(* Logix 5000 project; controller PLC_MCC1300_75F1 vendor 1 type 14 code 166 rev 32.11; software revision 32.04; part 53 of 83 *)
(* tags used below, declared in another part *)
   AUX_tConvoy_SL_NULL : UDT_Convoy_SL;
   AUX_xInitialize : BOOL;
   CONST_rgdDestMask : DINT[32];   // Destination Mask
   CONST_tPlant : UDT_PLANT_CONSTANTS;
   GP_TrackingGetFirstPlateInConveyor : GP_TrackingGetFirstPlateInConveyor;
   GP_TrackingPresencePlate : GP_TrackingPresencePlate;
   GP_TrackingSearchPlate : GP_TrackingSearchPlate;
   M310_M1_DR_R1 : AXIS_CIP_DRIVE;
   M310_xReqStopPrevConvForPos : BOOL;
   M310Popup : MAC_Popup_ZC[2];
   M310Popup_ReentryCap : UDT_ConvoyCap_ZC;
   M310Popup_SL_DATA : UDT_Convoy_SL;
   M310Popup_xDrivePosEnable : BOOL;
   M310Popup_xEndRise : BOOL;
   M310Popup_xEndRiseWaitingForCondition : BOOL;
   Sbr_INO_tConvoy_SL : UDT_Convoy_SL;
   TMP_d : DINT;
   TMP_dBaryc_ins_max : DINT;
   TMP_dBaryc_ins_min : DINT;
   TMP_dIndex : DINT;
   TMP_dIndex2 : DINT;
   TMP_dIndex3 : DINT;
   TMP_dStart0 : DINT;
   TMP_dStart1 : DINT;
   TMP_dStartSearchStop : DINT;
   TMP_dStop0 : DINT;
   TMP_dStop1 : DINT;
   TMP_dStopSearchStop : DINT;
   TMP_StartPlusLength : DINT;
   TMP_xAllCullet : BOOL;
   TMP_xAllLiteToCullet : BOOL;
   TMP_xAtLeastOneForSideLeg : BOOL;
   TMP_xPosHead : BOOL;
   TMP_xReqStopM310M1 : BOOL;
   TMP_xReqStopM310M2 : BOOL;
   TMP_xReqStopM310M3 : BOOL;
   xAlwaysOFF : BOOL;
   xDebugOFF : BOOL;
   Z300_BufferPlate : UDT_LINE_BUFFER_PLATE;
   Z300_Conveyor : UDT_StandConv[29];
   Z300_Conveyor_IN_MOTION : MAC_Conveyor_ZC_IN_MOTION[29];
   Z300_LineTracking : UDT_LINE_TRACKING;
   Z301 : MAC_Zone_ML;
(* MainProgram, continued *)

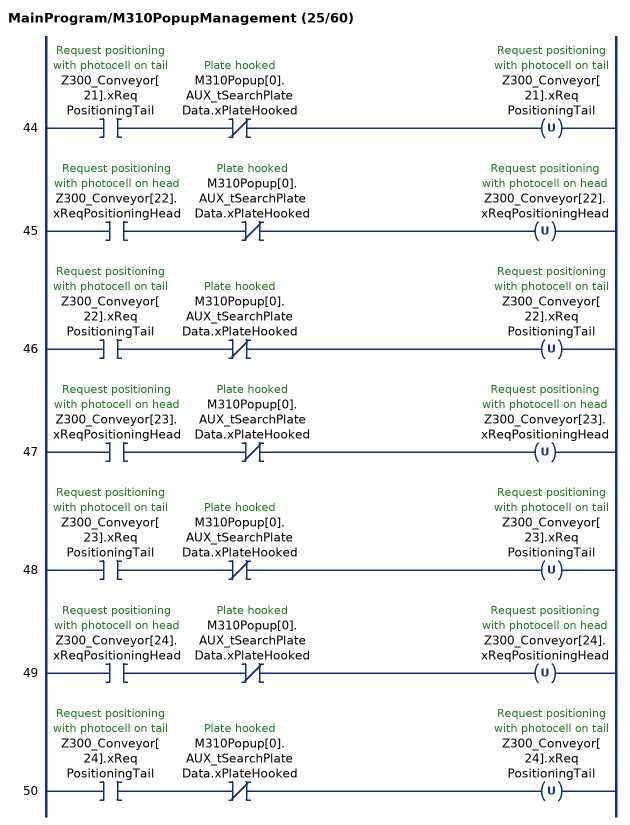
   [picture p841: MainProgram/M310PopupManagement rungs 44-50]
   44: XIC(Z300_Conveyor[21].xReqPositioningTail)XIO(M310Popup[0].AUX_tSearchPlateData.xPlateHooked)OTU(Z300_Conveyor[21].xReqPositioningTail);
   45: XIC(Z300_Conveyor[22].xReqPositioningHead)XIO(M310Popup[0].AUX_tSearchPlateData.xPlateHooked)OTU(Z300_Conveyor[22].xReqPositioningHead);
   46: XIC(Z300_Conveyor[22].xReqPositioningTail)XIO(M310Popup[0].AUX_tSearchPlateData.xPlateHooked)OTU(Z300_Conveyor[22].xReqPositioningTail);
   47: XIC(Z300_Conveyor[23].xReqPositioningHead)XIO(M310Popup[0].AUX_tSearchPlateData.xPlateHooked)OTU(Z300_Conveyor[23].xReqPositioningHead);
   48: XIC(Z300_Conveyor[23].xReqPositioningTail)XIO(M310Popup[0].AUX_tSearchPlateData.xPlateHooked)OTU(Z300_Conveyor[23].xReqPositioningTail);
   49: XIC(Z300_Conveyor[24].xReqPositioningHead)XIO(M310Popup[0].AUX_tSearchPlateData.xPlateHooked)OTU(Z300_Conveyor[24].xReqPositioningHead);
   50: XIC(Z300_Conveyor[24].xReqPositioningTail)XIO(M310Popup[0].AUX_tSearchPlateData.xPlateHooked)OTU(Z300_Conveyor[24].xReqPositioningTail);
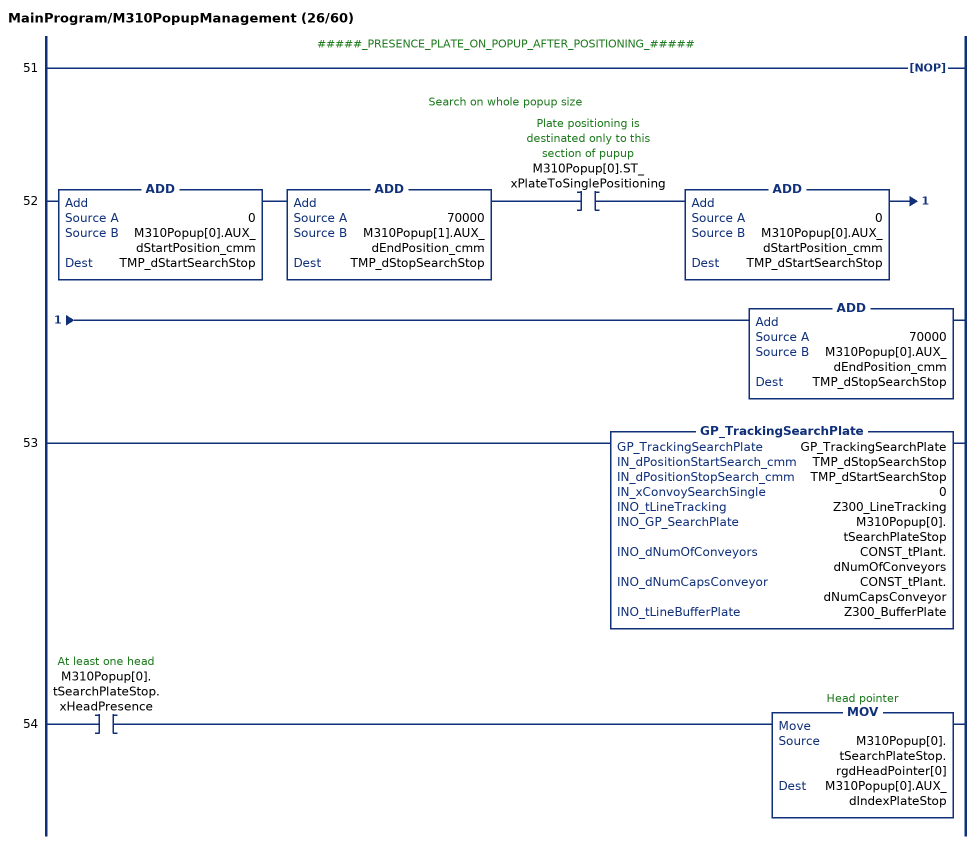
   // #####_PRESENCE_PLATE_ON_POPUP_AFTER_POSITIONING_#####
   51: NOP();
   // Search on whole popup size
   52: ADD(0,M310Popup[0].AUX_dStartPosition_cmm,TMP_dStartSearchStop)ADD(70000,M310Popup[1].AUX_dEndPosition_cmm,TMP_dStopSearchStop)XIC(M310Popup[0].ST_xPlateToSinglePositioning)ADD(0,M310Popup[0].AUX_dStartPosition_cmm,TMP_dStartSearchStop)ADD(70000,M310Popup[0].AUX_dEndPosition_cmm,TMP_dStopSearchStop);
   53: GP_TrackingSearchPlate(GP_TrackingSearchPlate,TMP_dStopSearchStop,TMP_dStartSearchStop,0,Z300_LineTracking,M310Popup[0].tSearchPlateStop,CONST_tPlant.dNumOfConveyors,CONST_tPlant.dNumCapsConveyor,Z300_BufferPlate);
   54: XIC(M310Popup[0].tSearchPlateStop.xHeadPresence)MOV(M310Popup[0].tSearchPlateStop.rgdHeadPointer[0],M310Popup[0].AUX_dIndexPlateStop);
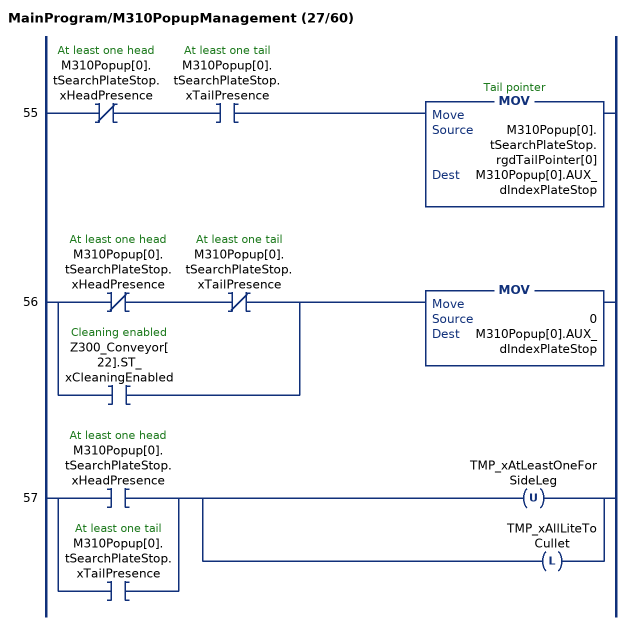
   55: XIO(M310Popup[0].tSearchPlateStop.xHeadPresence)XIC(M310Popup[0].tSearchPlateStop.xTailPresence)MOV(M310Popup[0].tSearchPlateStop.rgdTailPointer[0],M310Popup[0].AUX_dIndexPlateStop);
   56: [XIO(M310Popup[0].tSearchPlateStop.xHeadPresence) XIO(M310Popup[0].tSearchPlateStop.xTailPresence) ,XIC(Z300_Conveyor[22].ST_xCleaningEnabled) ]MOV(0,M310Popup[0].AUX_dIndexPlateStop);
   57: [XIC(M310Popup[0].tSearchPlateStop.xHeadPresence) ,XIC(M310Popup[0].tSearchPlateStop.xTailPresence) ][OTU(TMP_xAtLeastOneForSideLeg) ,OTL(TMP_xAllLiteToCullet) ];
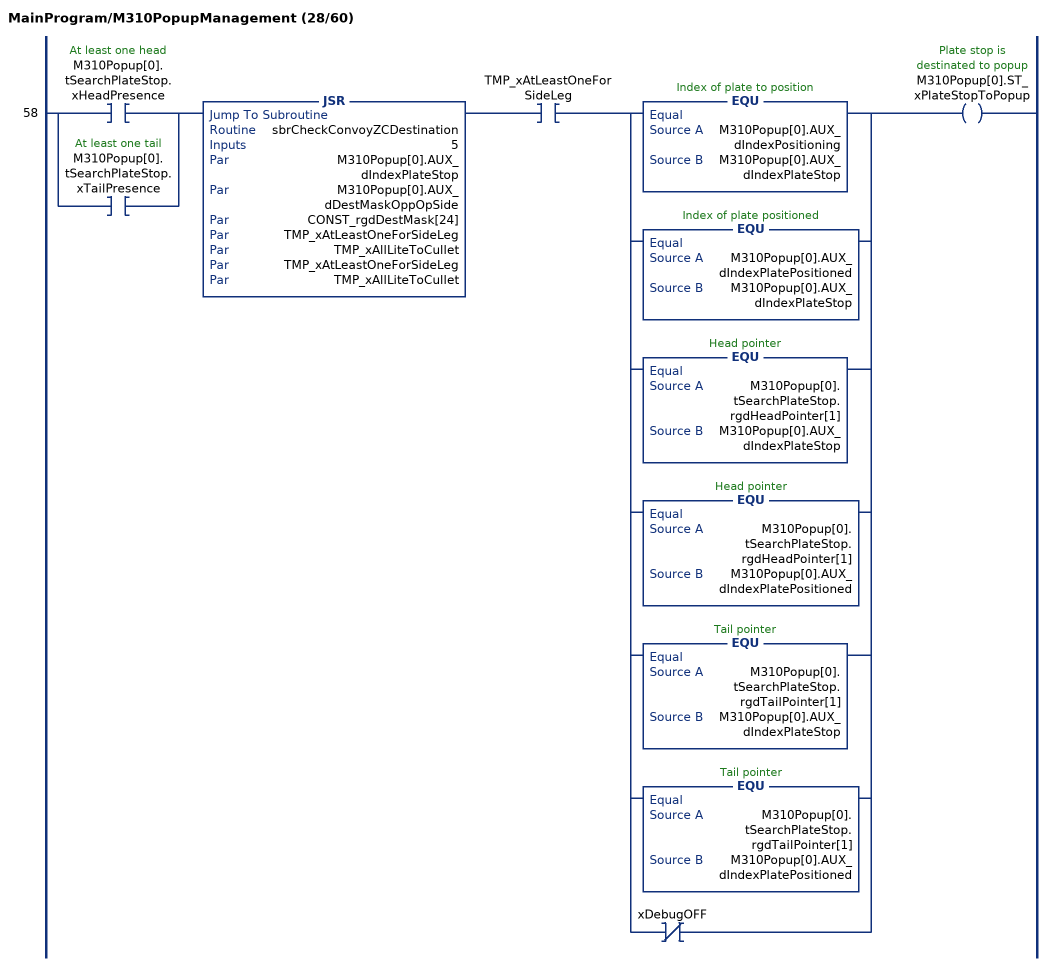
   58: [XIC(M310Popup[0].tSearchPlateStop.xHeadPresence) ,XIC(M310Popup[0].tSearchPlateStop.xTailPresence) ]JSR(sbrCheckConvoyZCDestination,5,M310Popup[0].AUX_dIndexPlateStop,M310Popup[0].AUX_dDestMaskOppOpSide,CONST_rgdDestMask[24],TMP_xAtLeastOneForSideLeg,TMP_xAllLiteToCullet,TMP_xAtLeastOneForSideLeg,TMP_xAllLiteToCullet)XIC(TMP_xAtLeastOneForSideLeg)[EQU(M310Popup[0].AUX_dIndexPositioning,M310Popup[0].AUX_dIndexPlateStop) ,EQU(M310Popup[0].AUX_dIndexPlatePositioned,M310Popup[0].AUX_dIndexPlateStop) ,EQU(M310Popup[0].tSearchPlateStop.rgdHeadPointer[1],M310Popup[0].AUX_dIndexPlateStop) ,EQU(M310Popup[0].tSearchPlateStop.rgdHeadPointer[1],M310Popup[0].AUX_dIndexPlatePositioned) ,EQU(M310Popup[0].tSearchPlateStop.rgdTailPointer[1],M310Popup[0].AUX_dIndexPlateStop) ,EQU(M310Popup[0].tSearchPlateStop.rgdTailPointer[1],M310Popup[0].AUX_dIndexPlatePositioned) ,XIO(xDebugOFF) ]OTE(M310Popup[0].ST_xPlateStopToPopup);
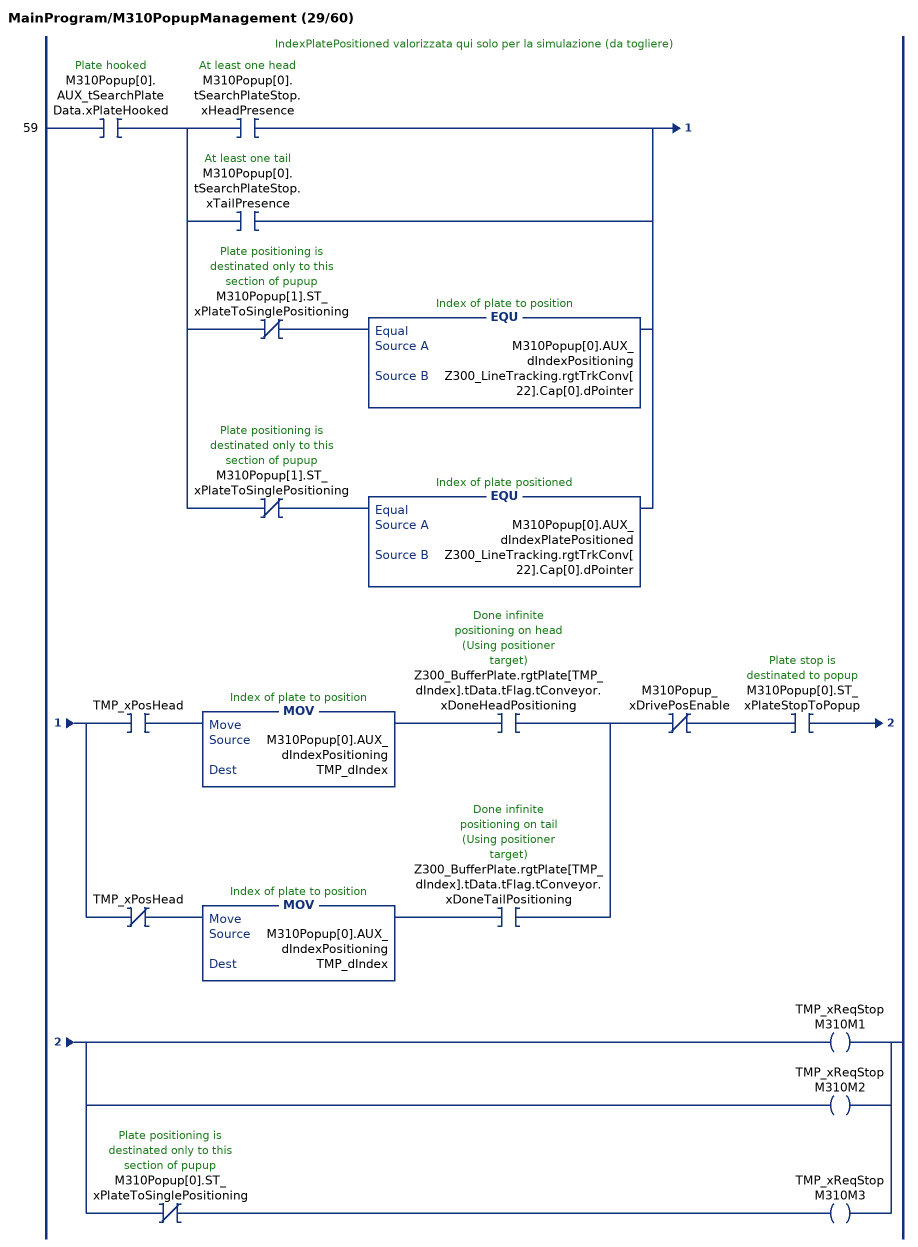
   // IndexPlatePositioned valorizzata qui solo per la simulazione (da togliere)
   59: XIC(M310Popup[0].AUX_tSearchPlateData.xPlateHooked)[XIC(M310Popup[0].tSearchPlateStop.xHeadPresence) ,XIC(M310Popup[0].tSearchPlateStop.xTailPresence) ,XIO(M310Popup[1].ST_xPlateToSinglePositioning) EQU(M310Popup[0].AUX_dIndexPositioning,Z300_LineTracking.rgtTrkConv[22].Cap[0].dPointer) ,XIO(M310Popup[1].ST_xPlateToSinglePositioning) EQU(M310Popup[0].AUX_dIndexPlatePositioned,Z300_LineTracking.rgtTrkConv[22].Cap[0].dPointer) ][XIC(TMP_xPosHead) MOV(M310Popup[0].AUX_dIndexPositioning,TMP_dIndex) XIC(Z300_BufferPlate.rgtPlate[TMP_dIndex].tData.tFlag.tConveyor.xDoneHeadPositioning) ,XIO(TMP_xPosHead) MOV(M310Popup[0].AUX_dIndexPositioning,TMP_dIndex) XIC(Z300_BufferPlate.rgtPlate[TMP_dIndex].tData.tFlag.tConveyor.xDoneTailPositioning) ]XIO(M310Popup_xDrivePosEnable)XIC(M310Popup[0].ST_xPlateStopToPopup)[OTE(TMP_xReqStopM310M1) ,OTE(TMP_xReqStopM310M2) ,XIO(M310Popup[0].ST_xPlateToSinglePositioning) OTE(TMP_xReqStopM310M3) ];
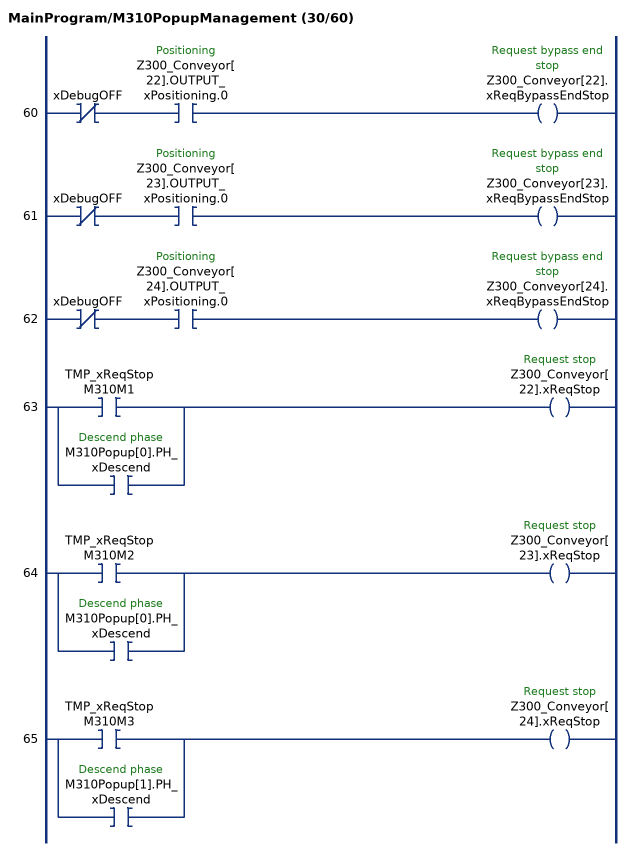
   60: XIO(xDebugOFF)XIC(Z300_Conveyor[22].OUTPUT_xPositioning.0)OTE(Z300_Conveyor[22].xReqBypassEndStop);
   61: XIO(xDebugOFF)XIC(Z300_Conveyor[23].OUTPUT_xPositioning.0)OTE(Z300_Conveyor[23].xReqBypassEndStop);
   62: XIO(xDebugOFF)XIC(Z300_Conveyor[24].OUTPUT_xPositioning.0)OTE(Z300_Conveyor[24].xReqBypassEndStop);
   63: [XIC(TMP_xReqStopM310M1) ,XIC(M310Popup[0].PH_xDescend) ]OTE(Z300_Conveyor[22].xReqStop);
   64: [XIC(TMP_xReqStopM310M2) ,XIC(M310Popup[0].PH_xDescend) ]OTE(Z300_Conveyor[23].xReqStop);
   65: [XIC(TMP_xReqStopM310M3) ,XIC(M310Popup[1].PH_xDescend) ]OTE(Z300_Conveyor[24].xReqStop);
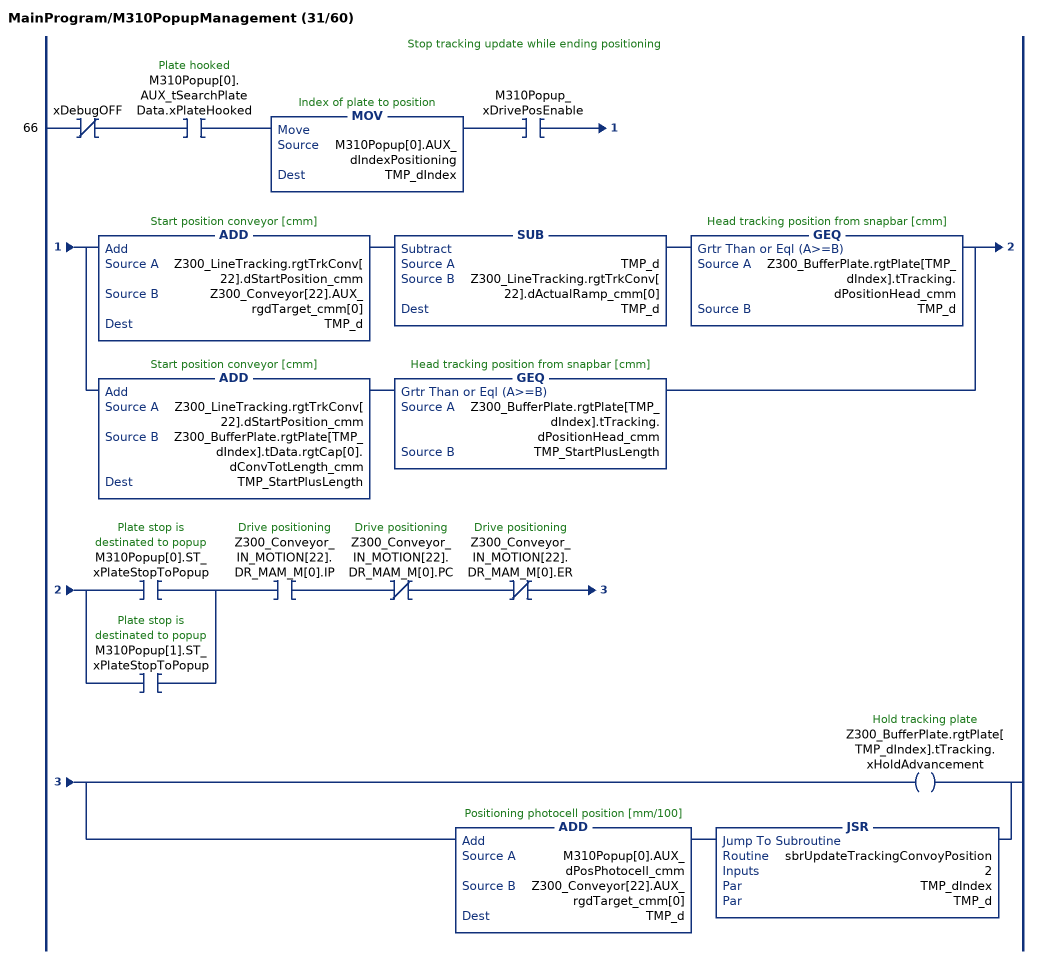
   // Stop tracking update while ending positioning
   66: XIO(xDebugOFF)XIC(M310Popup[0].AUX_tSearchPlateData.xPlateHooked)MOV(M310Popup[0].AUX_dIndexPositioning,TMP_dIndex)XIC(M310Popup_xDrivePosEnable)[ADD(Z300_LineTracking.rgtTrkConv[22].dStartPosition_cmm,Z300_Conveyor[22].AUX_rgdTarget_cmm[0],TMP_d) SUB(TMP_d,Z300_LineTracking.rgtTrkConv[22].dActualRamp_cmm[0],TMP_d) GEQ(Z300_BufferPlate.rgtPlate[TMP_dIndex].tTracking.dPositionHead_cmm,TMP_d) ,ADD(Z300_LineTracking.rgtTrkConv[22].dStartPosition_cmm,Z300_BufferPlate.rgtPlate[TMP_dIndex].tData.rgtCap[0].dConvTotLength_cmm,TMP_StartPlusLength) GEQ(Z300_BufferPlate.rgtPlate[TMP_dIndex].tTracking.dPositionHead_cmm,TMP_StartPlusLength) ][XIC(M310Popup[0].ST_xPlateStopToPopup) ,XIC(M310Popup[1].ST_xPlateStopToPopup) ]XIC(Z300_Conveyor_IN_MOTION[22].DR_MAM_M[0].IP)XIO(Z300_Conveyor_IN_MOTION[22].DR_MAM_M[0].PC)XIO(Z300_Conveyor_IN_MOTION[22].DR_MAM_M[0].ER)[OTE(Z300_BufferPlate.rgtPlate[TMP_dIndex].tTracking.xHoldAdvancement) ,ADD(M310Popup[0].AUX_dPosPhotocell_cmm,Z300_Conveyor[22].AUX_rgdTarget_cmm[0],TMP_d) JSR(sbrUpdateTrackingConvoyPosition,2,TMP_dIndex,TMP_d) ];
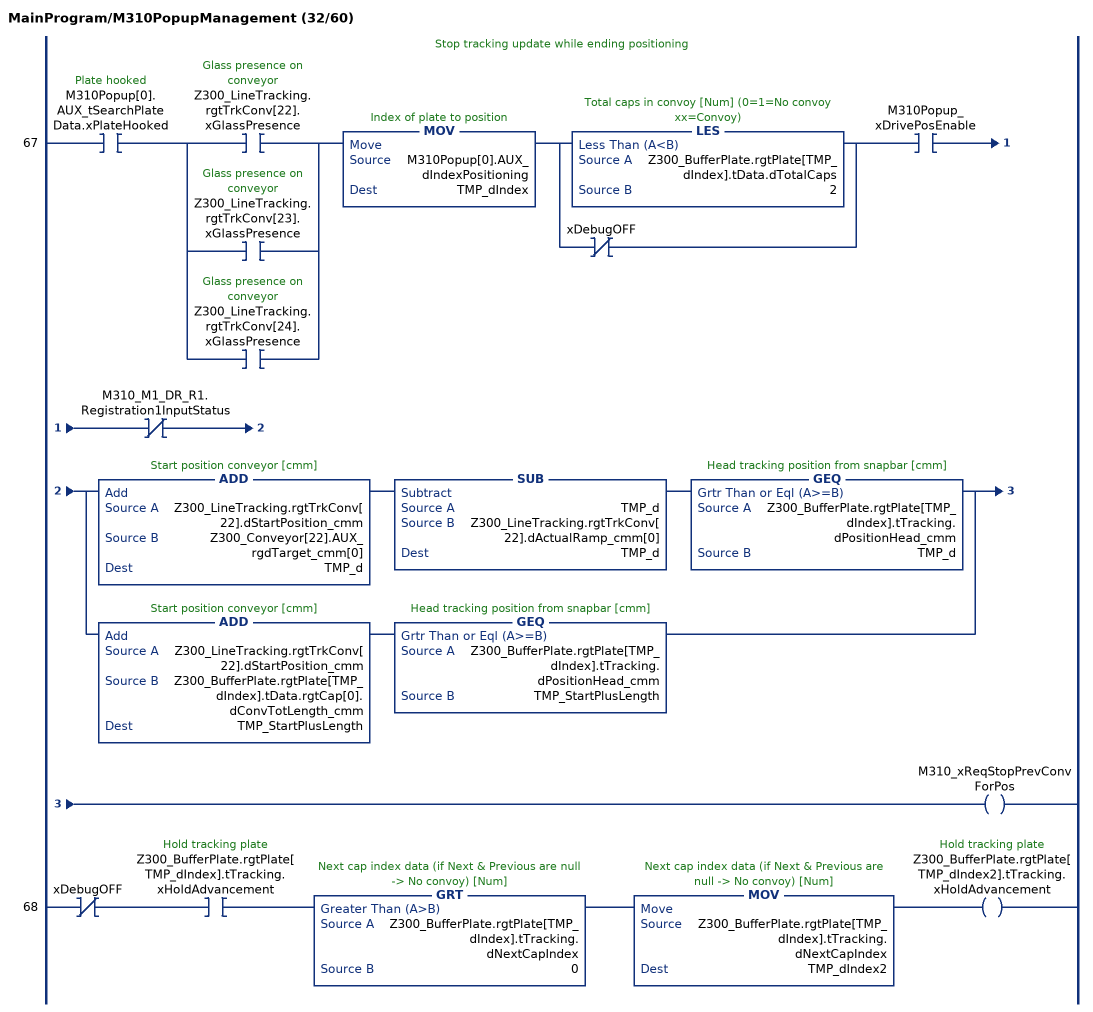
   // Stop tracking update while ending positioning
   67: XIC(M310Popup[0].AUX_tSearchPlateData.xPlateHooked)[XIC(Z300_LineTracking.rgtTrkConv[22].xGlassPresence) ,XIC(Z300_LineTracking.rgtTrkConv[23].xGlassPresence) ,XIC(Z300_LineTracking.rgtTrkConv[24].xGlassPresence) ]MOV(M310Popup[0].AUX_dIndexPositioning,TMP_dIndex)[LES(Z300_BufferPlate.rgtPlate[TMP_dIndex].tData.dTotalCaps,2) ,XIO(xDebugOFF) ]XIC(M310Popup_xDrivePosEnable)XIO(M310_M1_DR_R1.Registration1InputStatus)[ADD(Z300_LineTracking.rgtTrkConv[22].dStartPosition_cmm,Z300_Conveyor[22].AUX_rgdTarget_cmm[0],TMP_d) SUB(TMP_d,Z300_LineTracking.rgtTrkConv[22].dActualRamp_cmm[0],TMP_d) GEQ(Z300_BufferPlate.rgtPlate[TMP_dIndex].tTracking.dPositionHead_cmm,TMP_d) ,ADD(Z300_LineTracking.rgtTrkConv[22].dStartPosition_cmm,Z300_BufferPlate.rgtPlate[TMP_dIndex].tData.rgtCap[0].dConvTotLength_cmm,TMP_StartPlusLength) GEQ(Z300_BufferPlate.rgtPlate[TMP_dIndex].tTracking.dPositionHead_cmm,TMP_StartPlusLength) ]OTE(M310_xReqStopPrevConvForPos);
   68: XIO(xDebugOFF)XIC(Z300_BufferPlate.rgtPlate[TMP_dIndex].tTracking.xHoldAdvancement)GRT(Z300_BufferPlate.rgtPlate[TMP_dIndex].tTracking.dNextCapIndex,0)MOV(Z300_BufferPlate.rgtPlate[TMP_dIndex].tTracking.dNextCapIndex,TMP_dIndex2)OTE(Z300_BufferPlate.rgtPlate[TMP_dIndex2].tTracking.xHoldAdvancement);
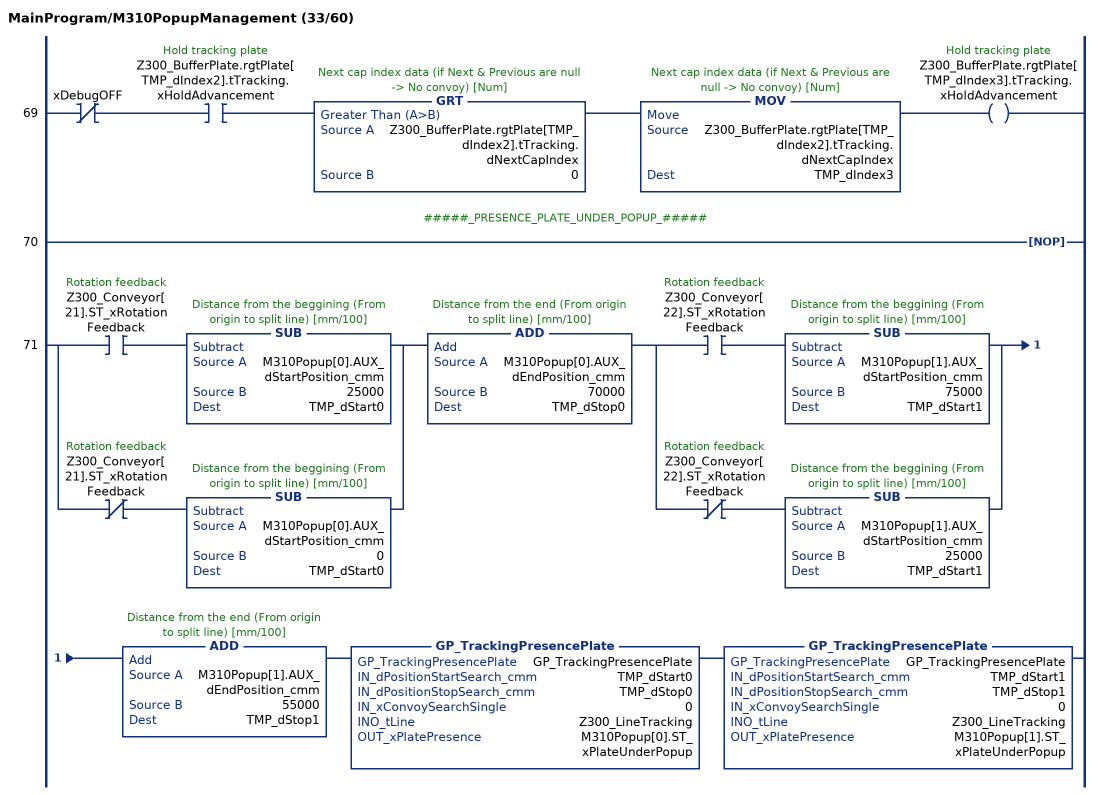
   69: XIO(xDebugOFF)XIC(Z300_BufferPlate.rgtPlate[TMP_dIndex2].tTracking.xHoldAdvancement)GRT(Z300_BufferPlate.rgtPlate[TMP_dIndex2].tTracking.dNextCapIndex,0)MOV(Z300_BufferPlate.rgtPlate[TMP_dIndex2].tTracking.dNextCapIndex,TMP_dIndex3)OTE(Z300_BufferPlate.rgtPlate[TMP_dIndex3].tTracking.xHoldAdvancement);
   // #####_PRESENCE_PLATE_UNDER_POPUP_#####
   70: NOP();
   71: [XIC(Z300_Conveyor[21].ST_xRotationFeedback) SUB(M310Popup[0].AUX_dStartPosition_cmm,25000,TMP_dStart0) ,XIO(Z300_Conveyor[21].ST_xRotationFeedback) SUB(M310Popup[0].AUX_dStartPosition_cmm,0,TMP_dStart0) ]ADD(M310Popup[0].AUX_dEndPosition_cmm,70000,TMP_dStop0)[XIC(Z300_Conveyor[22].ST_xRotationFeedback) SUB(M310Popup[1].AUX_dStartPosition_cmm,75000,TMP_dStart1) ,XIO(Z300_Conveyor[22].ST_xRotationFeedback) SUB(M310Popup[1].AUX_dStartPosition_cmm,25000,TMP_dStart1) ]ADD(M310Popup[1].AUX_dEndPosition_cmm,55000,TMP_dStop1)GP_TrackingPresencePlate(GP_TrackingPresencePlate,TMP_dStart0,TMP_dStop0,0,Z300_LineTracking,M310Popup[0].ST_xPlateUnderPopup)GP_TrackingPresencePlate(GP_TrackingPresencePlate,TMP_dStart1,TMP_dStop1,0,Z300_LineTracking,M310Popup[1].ST_xPlateUnderPopup);
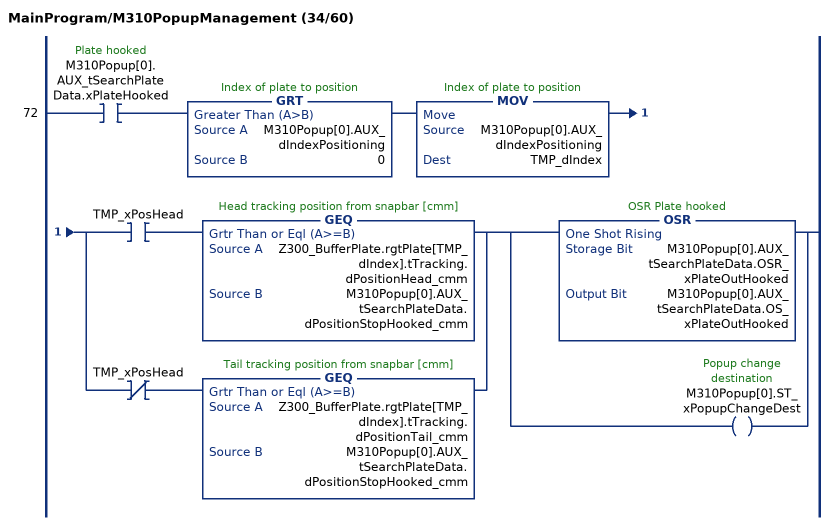
   72: XIC(M310Popup[0].AUX_tSearchPlateData.xPlateHooked)GRT(M310Popup[0].AUX_dIndexPositioning,0)MOV(M310Popup[0].AUX_dIndexPositioning,TMP_dIndex)[XIC(TMP_xPosHead) GEQ(Z300_BufferPlate.rgtPlate[TMP_dIndex].tTracking.dPositionHead_cmm,M310Popup[0].AUX_tSearchPlateData.dPositionStopHooked_cmm) ,XIO(TMP_xPosHead) GEQ(Z300_BufferPlate.rgtPlate[TMP_dIndex].tTracking.dPositionTail_cmm,M310Popup[0].AUX_tSearchPlateData.dPositionStopHooked_cmm) ][OSR(M310Popup[0].AUX_tSearchPlateData.OSR_xPlateOutHooked,M310Popup[0].AUX_tSearchPlateData.OS_xPlateOutHooked) ,OTE(M310Popup[0].ST_xPopupChangeDest) ];
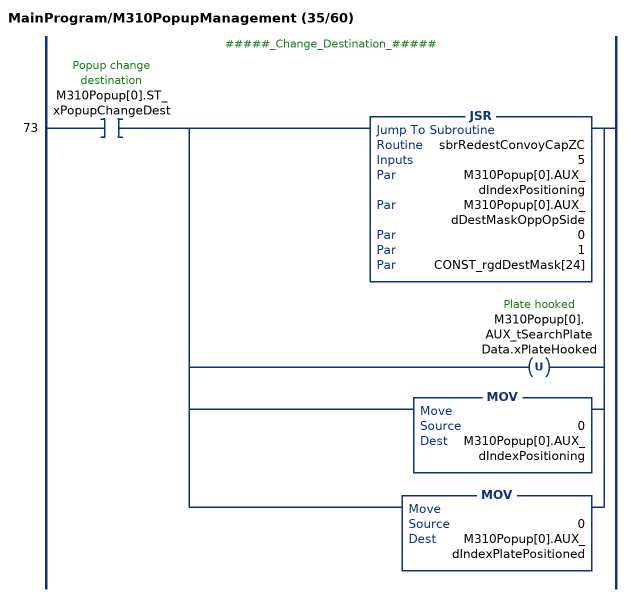
   // #####_Change_Destination_#####
   73: XIC(M310Popup[0].ST_xPopupChangeDest)[JSR(sbrRedestConvoyCapZC,5,M310Popup[0].AUX_dIndexPositioning,M310Popup[0].AUX_dDestMaskOppOpSide,0,1,CONST_rgdDestMask[24]) ,OTU(M310Popup[0].AUX_tSearchPlateData.xPlateHooked) ,MOV(0,M310Popup[0].AUX_dIndexPositioning) ,MOV(0,M310Popup[0].AUX_dIndexPlatePositioned) ];